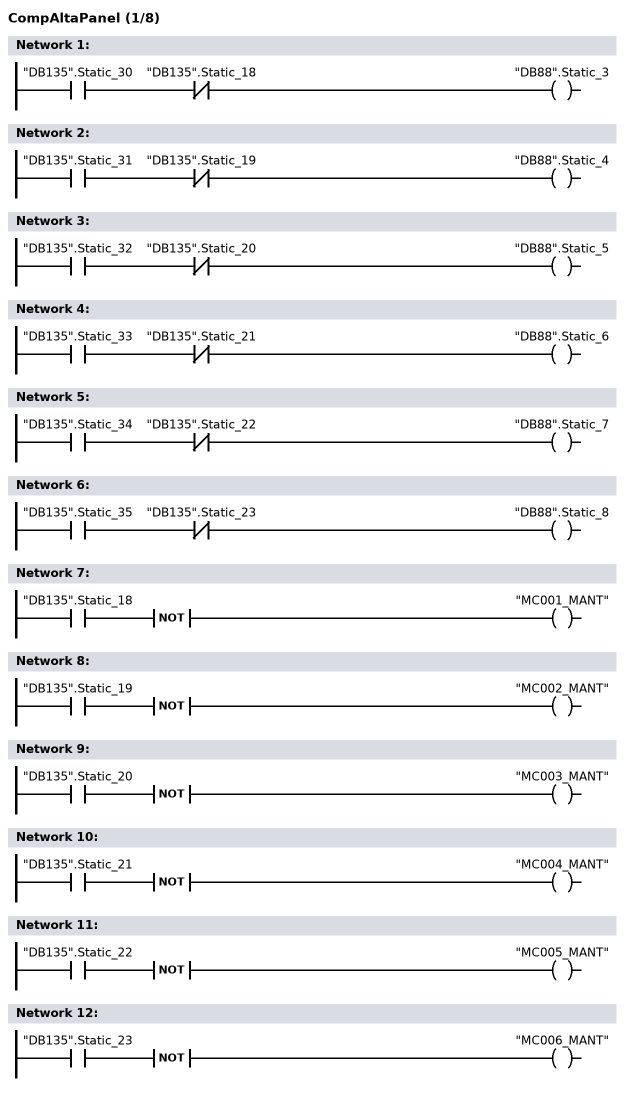
   RUNG wire#powerrail
      Contact( "DB135".Static_30 )
      I_Contact( "DB135".Static_18 )
      Coil( "DB88".Static_3 )
   END_RUNG
   // the same network as SCL:
   "DB88".Static_3 := "DB135".Static_30 AND NOT "DB135".Static_18;
END_REGION

REGION Network 2
   RUNG wire#powerrail
      Contact( "DB135".Static_31 )
      I_Contact( "DB135".Static_19 )
      Coil( "DB88".Static_4 )
   END_RUNG
   // the same network as SCL:
   "DB88".Static_4 := "DB135".Static_31 AND NOT "DB135".Static_19;
END_REGION

REGION Network 3
   RUNG wire#powerrail
      Contact( "DB135".Static_32 )
      I_Contact( "DB135".Static_20 )
      Coil( "DB88".Static_5 )
   END_RUNG
   // the same network as SCL:
   "DB88".Static_5 := "DB135".Static_32 AND NOT "DB135".Static_20;
END_REGION

REGION Network 4
   RUNG wire#powerrail
      Contact( "DB135".Static_33 )
      I_Contact( "DB135".Static_21 )
      Coil( "DB88".Static_6 )
   END_RUNG
   // the same network as SCL:
   "DB88".Static_6 := "DB135".Static_33 AND NOT "DB135".Static_21;
END_REGION

REGION Network 5
   RUNG wire#powerrail
      Contact( "DB135".Static_34 )
      I_Contact( "DB135".Static_22 )
      Coil( "DB88".Static_7 )
   END_RUNG
   // the same network as SCL:
   "DB88".Static_7 := "DB135".Static_34 AND NOT "DB135".Static_22;
END_REGION

REGION Network 6
   RUNG wire#powerrail
      Contact( "DB135".Static_35 )
      I_Contact( "DB135".Static_23 )
      Coil( "DB88".Static_8 )
   END_RUNG
   // the same network as SCL:
   "DB88".Static_8 := "DB135".Static_35 AND NOT "DB135".Static_23;
END_REGION

REGION Network 7
   RUNG wire#powerrail
      Contact( "DB135".Static_18 )
      Not()
      Coil( "MC001_MANT" )
   END_RUNG
   // the same network as SCL:
   "MC001_MANT" := NOT "DB135".Static_18;
END_REGION

REGION Network 8
   RUNG wire#powerrail
      Contact( "DB135".Static_19 )
      Not()
      Coil( "MC002_MANT" )
   END_RUNG
   // the same network as SCL:
   "MC002_MANT" := NOT "DB135".Static_19;
END_REGION

REGION Network 9
   RUNG wire#powerrail
      Contact( "DB135".Static_20 )
      Not()
      Coil( "MC003_MANT" )
   END_RUNG
   // the same network as SCL:
   "MC003_MANT" := NOT "DB135".Static_20;
END_REGION

REGION Network 10
   RUNG wire#powerrail
      Contact( "DB135".Static_21 )
      Not()
      Coil( "MC004_MANT" )
   END_RUNG
   // the same network as SCL:
   "MC004_MANT" := NOT "DB135".Static_21;
END_REGION

REGION Network 11
   RUNG wire#powerrail
      Contact( "DB135".Static_22 )
      Not()
      Coil( "MC005_MANT" )
   END_RUNG
   // the same network as SCL:
   "MC005_MANT" := NOT "DB135".Static_22;
END_REGION

REGION Network 12
   RUNG wire#powerrail
      Contact( "DB135".Static_23 )
      Not()
      Coil( "MC006_MANT" )
   END_RUNG
   // the same network as SCL:
   "MC006_MANT" := NOT "DB135".Static_23;
END_REGION

REGION Network 13
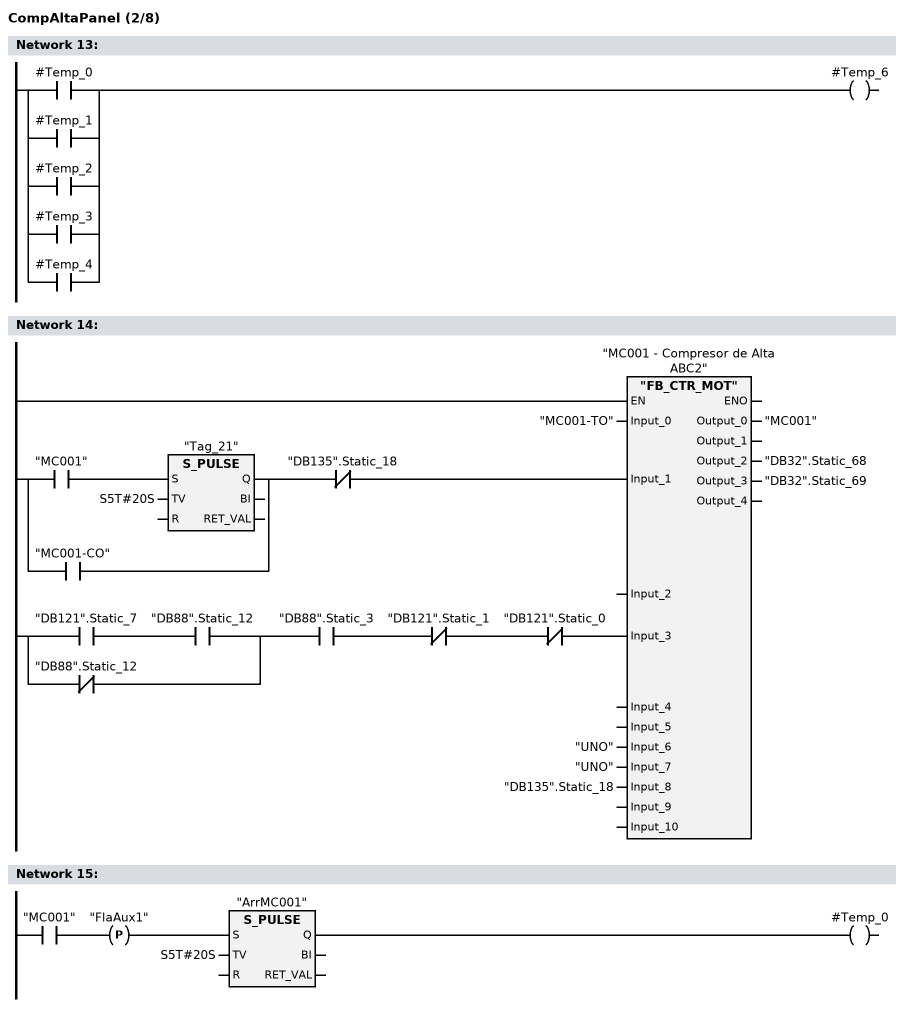
   RUNG wire#powerrail
      Contact( #Temp_0 )
      wire#w1
      Coil( #Temp_6 )
   END_RUNG
   RUNG wire#powerrail
      Contact( #Temp_1 )
   END_RUNG wire#w1
   RUNG wire#powerrail
      Contact( #Temp_2 )
   END_RUNG wire#w1
   RUNG wire#powerrail
      Contact( #Temp_3 )
   END_RUNG wire#w1
   RUNG wire#powerrail
      Contact( #Temp_4 )
   END_RUNG wire#w1
   // the same network as SCL:
   #Temp_6 := #Temp_0 OR #Temp_1 OR #Temp_2 OR #Temp_3 OR #Temp_4;
END_REGION

REGION Network 14
   #_s5time1 := S_PULSE(T_NO := "Tag_21", TV := S5T#20S, S := "MC001", Q => #_w1);
   "MC001 - Compresor de Alta ABC2"(Input_0 := "MC001-TO",   // "FB_CTR_MOT"
                           Input_1 := (#_w1 OR "MC001-CO") AND NOT "DB135".Static_18,
                           Input_3 := (("DB121".Static_7 AND "DB88".Static_12) OR NOT "DB88".Static_12) AND "DB88".Static_3 AND NOT "DB121".Static_1 AND NOT "DB121".Static_0,
                           Input_6 := "UNO",
                           Input_7 := "UNO",
                           Input_8 := "DB135".Static_18,
                           Output_0 => "MC001",
                           Output_2 => "DB32".Static_68,
                           Output_3 => "DB32".Static_69);
END_REGION

REGION Network 15
   RUNG wire#powerrail
      Contact( "MC001" )
      P_Trig( "FlaAux1" )
      S_PULSE(T_NO := "ArrMC001", TV := S5T#20S, R :=, BI =>, RET_VAL =>)
      Coil( #Temp_0 )
   END_RUNG
   // the same network as SCL:
   #_w1 := "MC001" AND NOT "FlaAux1";   // rising edge
   "FlaAux1" := "MC001";
   #_s5time1 := S_PULSE(T_NO := "ArrMC001", S := #_w1, TV := S5T#20S, Q => #_w2);
   #Temp_0 := #_w2;
END_REGION

REGION Network 16
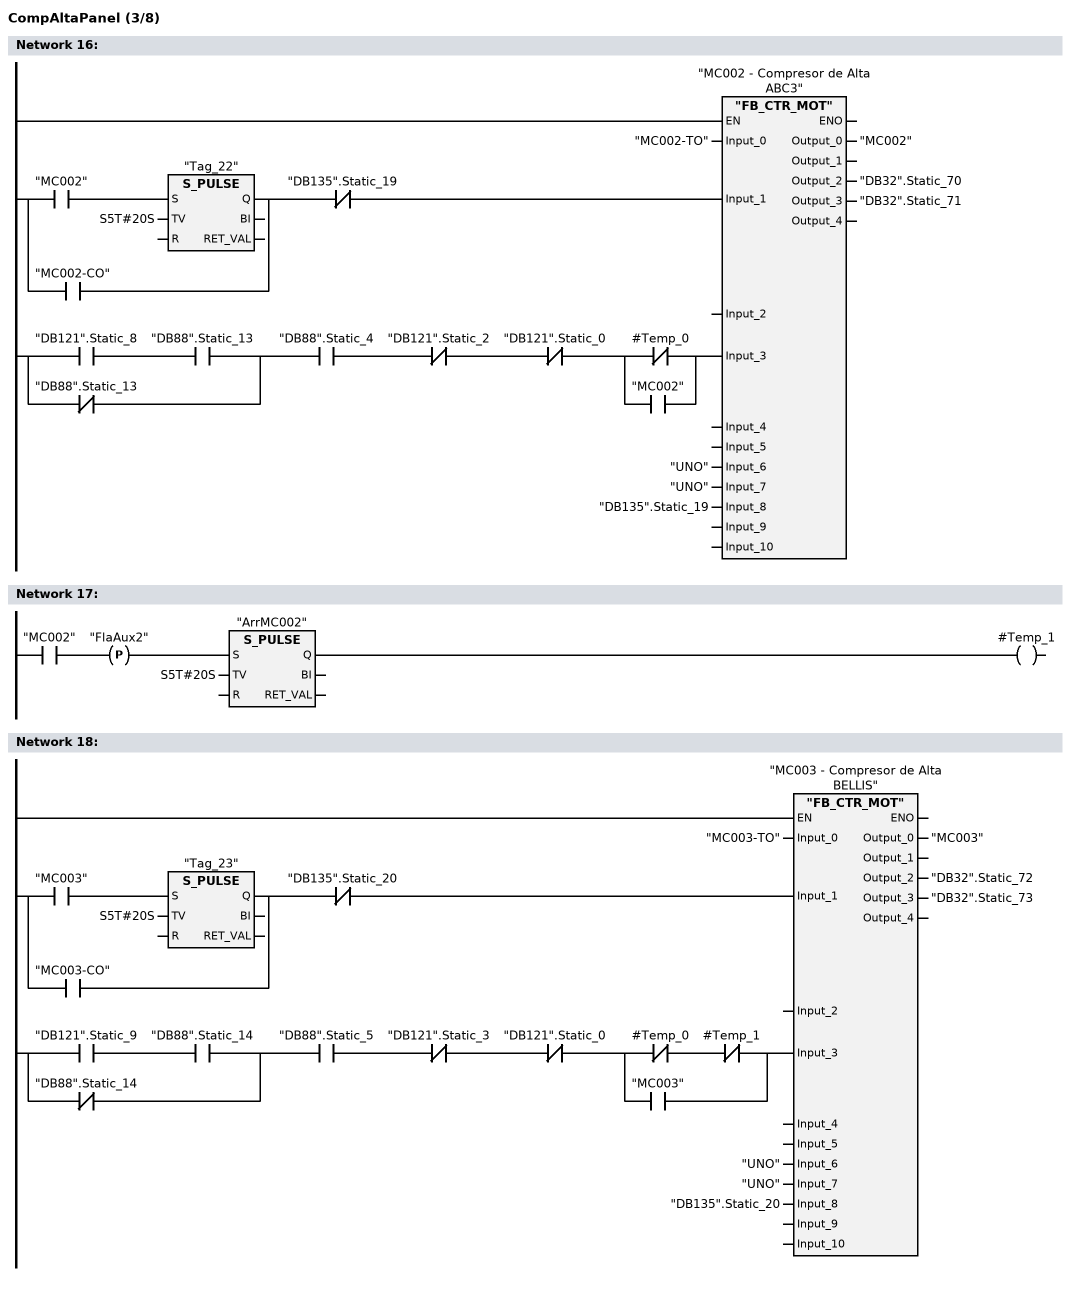
   #_s5time1 := S_PULSE(T_NO := "Tag_22", TV := S5T#20S, S := "MC002", Q => #_w1);
   "MC002 - Compresor de Alta ABC3"(Input_0 := "MC002-TO",   // "FB_CTR_MOT"
                           Input_1 := (#_w1 OR "MC002-CO") AND NOT "DB135".Static_19,
                           Input_3 := (("DB121".Static_8 AND "DB88".Static_13) OR NOT "DB88".Static_13) AND "DB88".Static_4 AND NOT "DB121".Static_2 AND NOT "DB121".Static_0 AND (NOT #Temp_0 OR "MC002"),
                           Input_6 := "UNO",
                           Input_7 := "UNO",
                           Input_8 := "DB135".Static_19,
                           Output_0 => "MC002",
                           Output_2 => "DB32".Static_70,
                           Output_3 => "DB32".Static_71);
END_REGION

REGION Network 17
   RUNG wire#powerrail
      Contact( "MC002" )
      P_Trig( "FlaAux2" )
      S_PULSE(T_NO := "ArrMC002", TV := S5T#20S, R :=, BI =>, RET_VAL =>)
      Coil( #Temp_1 )
   END_RUNG
   // the same network as SCL:
   #_w1 := "MC002" AND NOT "FlaAux2";   // rising edge
   "FlaAux2" := "MC002";
   #_s5time1 := S_PULSE(T_NO := "ArrMC002", S := #_w1, TV := S5T#20S, Q => #_w2);
   #Temp_1 := #_w2;
END_REGION

REGION Network 18
   #_s5time1 := S_PULSE(T_NO := "Tag_23", TV := S5T#20S, S := "MC003", Q => #_w1);
   "MC003 - Compresor de Alta BELLIS"(Input_0 := "MC003-TO",   // "FB_CTR_MOT"
                           Input_1 := (#_w1 OR "MC003-CO") AND NOT "DB135".Static_20,
                           Input_3 := (("DB121".Static_9 AND "DB88".Static_14) OR NOT "DB88".Static_14) AND "DB88".Static_5 AND NOT "DB121".Static_3 AND NOT "DB121".Static_0 AND ((NOT #Temp_0 AND NOT #Temp_1) OR "MC003"),
                           Input_6 := "UNO",
                           Input_7 := "UNO",
                           Input_8 := "DB135".Static_20,
                           Output_0 => "MC003",
                           Output_2 => "DB32".Static_72,
                           Output_3 => "DB32".Static_73);
END_REGION

REGION Network 19
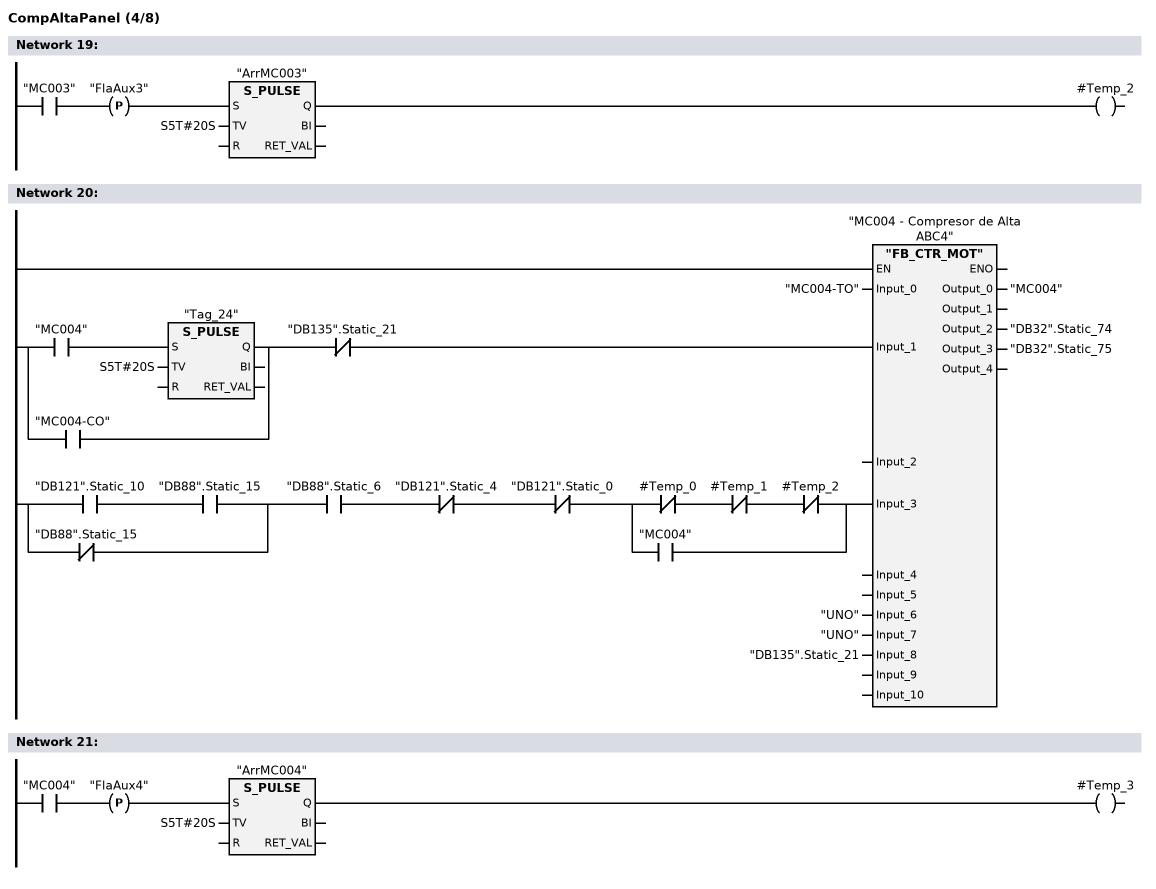
   RUNG wire#powerrail
      Contact( "MC003" )
      P_Trig( "FlaAux3" )
      S_PULSE(T_NO := "ArrMC003", TV := S5T#20S, R :=, BI =>, RET_VAL =>)
      Coil( #Temp_2 )
   END_RUNG
   // the same network as SCL:
   #_w1 := "MC003" AND NOT "FlaAux3";   // rising edge
   "FlaAux3" := "MC003";
   #_s5time1 := S_PULSE(T_NO := "ArrMC003", S := #_w1, TV := S5T#20S, Q => #_w2);
   #Temp_2 := #_w2;
END_REGION

REGION Network 20
   #_s5time1 := S_PULSE(T_NO := "Tag_24", TV := S5T#20S, S := "MC004", Q => #_w1);
   "MC004 - Compresor de Alta ABC4"(Input_0 := "MC004-TO",   // "FB_CTR_MOT"
                           Input_1 := (#_w1 OR "MC004-CO") AND NOT "DB135".Static_21,
                           Input_3 := (("DB121".Static_10 AND "DB88".Static_15) OR NOT "DB88".Static_15) AND "DB88".Static_6 AND NOT "DB121".Static_4 AND NOT "DB121".Static_0 AND ((NOT #Temp_0 AND NOT #Temp_1 AND NOT #Temp_2) OR "MC004"),
                           Input_6 := "UNO",
                           Input_7 := "UNO",
                           Input_8 := "DB135".Static_21,
                           Output_0 => "MC004",
                           Output_2 => "DB32".Static_74,
                           Output_3 => "DB32".Static_75);
END_REGION

REGION Network 21
   RUNG wire#powerrail
      Contact( "MC004" )
      P_Trig( "FlaAux4" )
      S_PULSE(T_NO := "ArrMC004", TV := S5T#20S, R :=, BI =>, RET_VAL =>)
      Coil( #Temp_3 )
   END_RUNG
   // the same network as SCL:
   #_w1 := "MC004" AND NOT "FlaAux4";   // rising edge
   "FlaAux4" := "MC004";
   #_s5time1 := S_PULSE(T_NO := "ArrMC004", S := #_w1, TV := S5T#20S, Q => #_w2);
   #Temp_3 := #_w2;
END_REGION

REGION Network 22
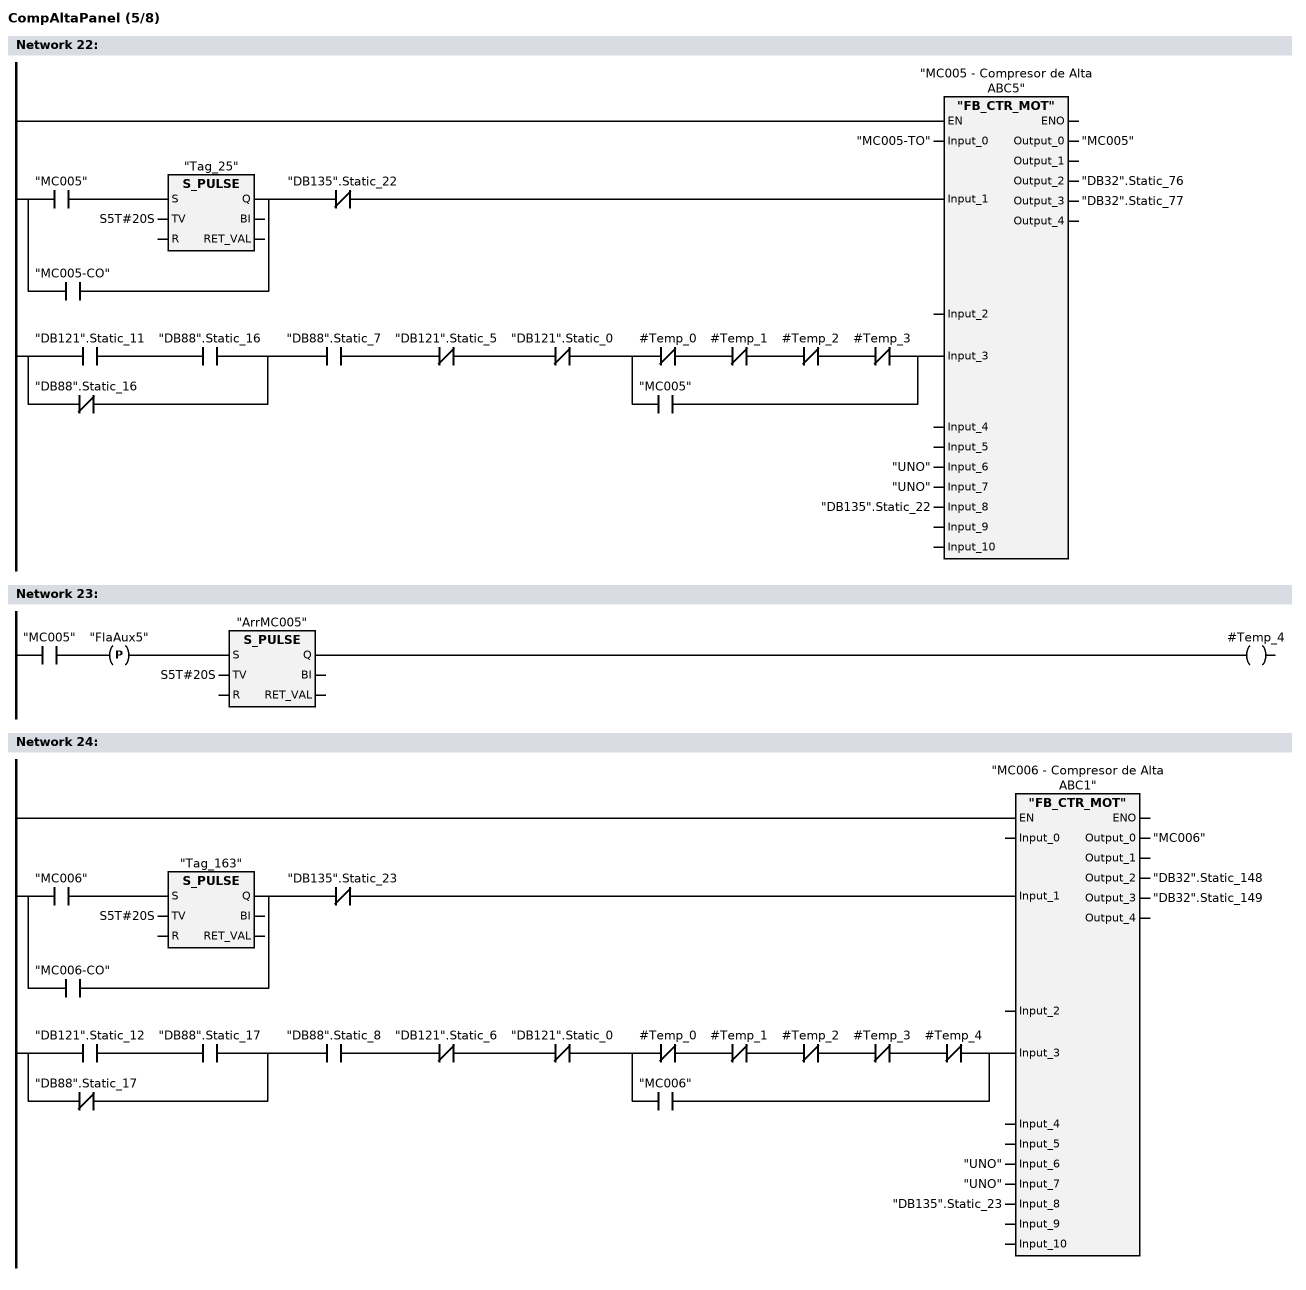
   #_s5time1 := S_PULSE(T_NO := "Tag_25", TV := S5T#20S, S := "MC005", Q => #_w1);
   "MC005 - Compresor de Alta ABC5"(Input_0 := "MC005-TO",   // "FB_CTR_MOT"
                           Input_1 := (#_w1 OR "MC005-CO") AND NOT "DB135".Static_22,
                           Input_3 := (("DB121".Static_11 AND "DB88".Static_16) OR NOT "DB88".Static_16) AND "DB88".Static_7 AND NOT "DB121".Static_5 AND NOT "DB121".Static_0 AND ((NOT #Temp_0 AND NOT #Temp_1 AND NOT #Temp_2 AND NOT #Temp_3) OR "MC005"),
                           Input_6 := "UNO",
                           Input_7 := "UNO",
                           Input_8 := "DB135".Static_22,
                           Output_0 => "MC005",
                           Output_2 => "DB32".Static_76,
                           Output_3 => "DB32".Static_77);
END_REGION

REGION Network 23
   RUNG wire#powerrail
      Contact( "MC005" )
      P_Trig( "FlaAux5" )
      S_PULSE(T_NO := "ArrMC005", TV := S5T#20S, R :=, BI =>, RET_VAL =>)
      Coil( #Temp_4 )
   END_RUNG
   // the same network as SCL:
   #_w1 := "MC005" AND NOT "FlaAux5";   // rising edge
   "FlaAux5" := "MC005";
   #_s5time1 := S_PULSE(T_NO := "ArrMC005", S := #_w1, TV := S5T#20S, Q => #_w2);
   #Temp_4 := #_w2;
END_REGION

REGION Network 24
   #_s5time1 := S_PULSE(T_NO := "Tag_163", TV := S5T#20S, S := "MC006", Q => #_w1);
   "MC006 - Compresor de Alta ABC1"(Input_1 := (#_w1 OR "MC006-CO") AND NOT "DB135".Static_23,   // "FB_CTR_MOT"
                           Input_3 := (("DB121".Static_12 AND "DB88".Static_17) OR NOT "DB88".Static_17) AND "DB88".Static_8 AND NOT "DB121".Static_6 AND NOT "DB121".Static_0 AND ((NOT #Temp_0 AND NOT #Temp_1 AND NOT #Temp_2 AND NOT #Temp_3 AND NOT #Temp_4) OR "MC006"),
                           Input_6 := "UNO",
                           Input_7 := "UNO",
                           Input_8 := "DB135".Static_23,
                           Output_0 => "MC006",
                           Output_2 => "DB32".Static_148,
                           Output_3 => "DB32".Static_149);
END_REGION

REGION Network 25
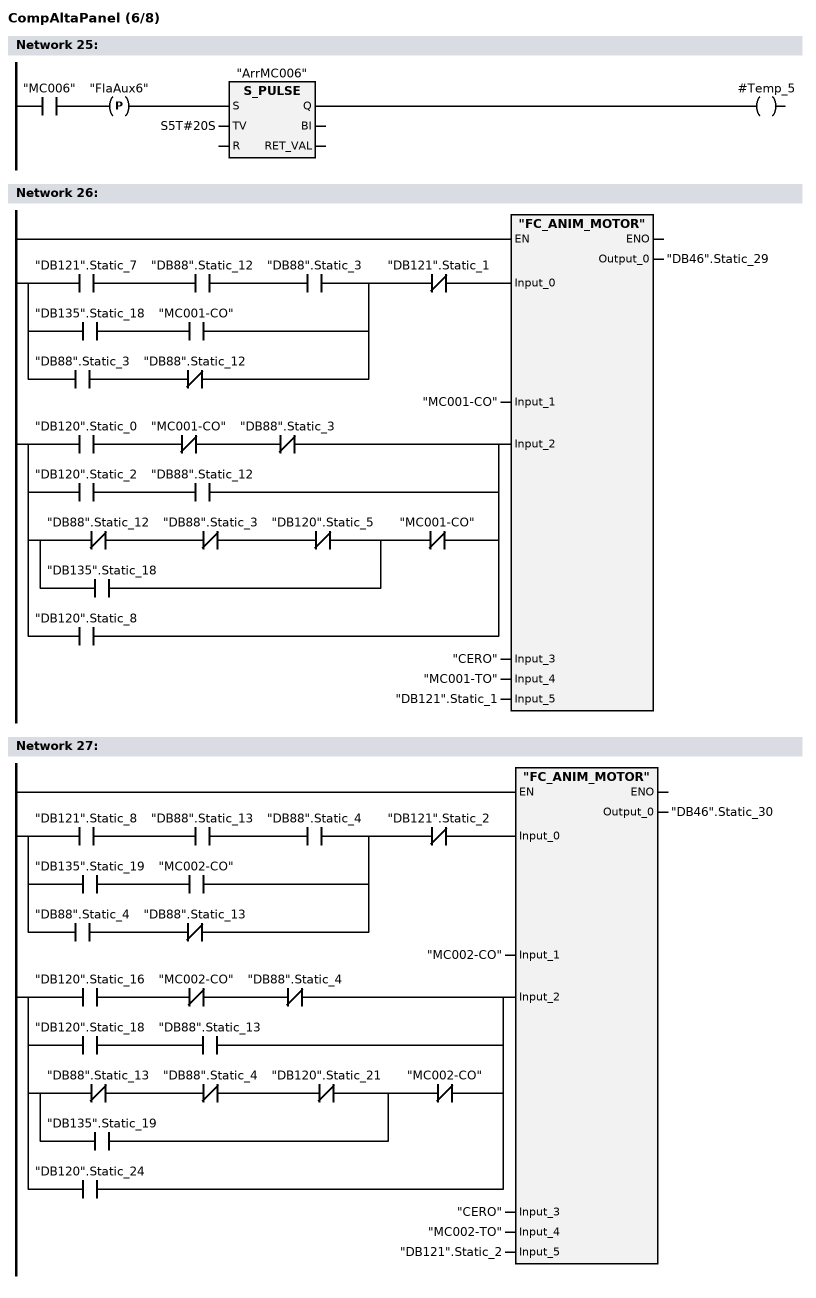
   RUNG wire#powerrail
      Contact( "MC006" )
      P_Trig( "FlaAux6" )
      S_PULSE(T_NO := "ArrMC006", TV := S5T#20S, R :=, BI =>, RET_VAL =>)
      Coil( #Temp_5 )
   END_RUNG
   // the same network as SCL:
   #_w1 := "MC006" AND NOT "FlaAux6";   // rising edge
   "FlaAux6" := "MC006";
   #_s5time1 := S_PULSE(T_NO := "ArrMC006", S := #_w1, TV := S5T#20S, Q => #_w2);
   #Temp_5 := #_w2;
END_REGION

REGION Network 26
   "FC_ANIM_MOTOR"(Input_0 := (("DB121".Static_7 AND "DB88".Static_12 AND "DB88".Static_3) OR ("DB135".Static_18 AND "MC001-CO") OR ("DB88".Static_3 AND NOT "DB88".Static_12)) AND NOT "DB121".Static_1,
                   Input_1 := "MC001-CO",
                   Input_2 := ("DB120".Static_0 AND NOT "MC001-CO" AND NOT "DB88".Static_3) OR ("DB120".Static_2 AND "DB88".Static_12) OR "DB120".Static_8 OR (("DB135".Static_18 OR (NOT "DB88".Static_12 AND NOT "DB88".Static_3 AND NOT "DB120".Static_5)) AND NOT "MC001-CO"),
                   Input_3 := "CERO",
                   Input_4 := "MC001-TO",
                   Input_5 := "DB121".Static_1,
                   Output_0 => "DB46".Static_29);
END_REGION

REGION Network 27
   "FC_ANIM_MOTOR"(Input_0 := (("DB121".Static_8 AND "DB88".Static_13 AND "DB88".Static_4) OR ("DB135".Static_19 AND "MC002-CO") OR ("DB88".Static_4 AND NOT "DB88".Static_13)) AND NOT "DB121".Static_2,
                   Input_1 := "MC002-CO",
                   Input_2 := ("DB120".Static_16 AND NOT "MC002-CO" AND NOT "DB88".Static_4) OR ("DB120".Static_18 AND "DB88".Static_13) OR "DB120".Static_24 OR (("DB135".Static_19 OR (NOT "DB88".Static_13 AND NOT "DB88".Static_4 AND NOT "DB120".Static_21)) AND NOT "MC002-CO"),
                   Input_3 := "CERO",
                   Input_4 := "MC002-TO",
                   Input_5 := "DB121".Static_2,
                   Output_0 => "DB46".Static_30);
END_REGION

REGION Network 28
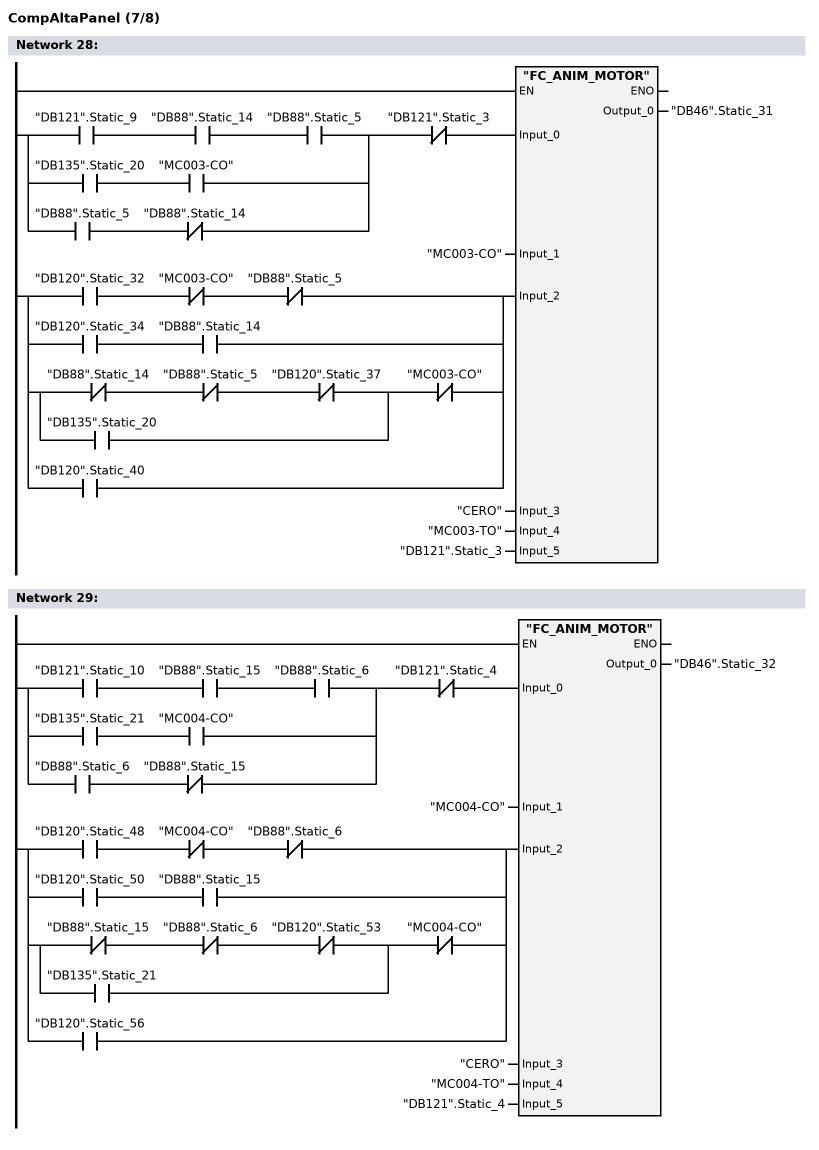
   "FC_ANIM_MOTOR"(Input_0 := (("DB121".Static_9 AND "DB88".Static_14 AND "DB88".Static_5) OR ("DB135".Static_20 AND "MC003-CO") OR ("DB88".Static_5 AND NOT "DB88".Static_14)) AND NOT "DB121".Static_3,
                   Input_1 := "MC003-CO",
                   Input_2 := ("DB120".Static_32 AND NOT "MC003-CO" AND NOT "DB88".Static_5) OR ("DB120".Static_34 AND "DB88".Static_14) OR "DB120".Static_40 OR (("DB135".Static_20 OR (NOT "DB88".Static_14 AND NOT "DB88".Static_5 AND NOT "DB120".Static_37)) AND NOT "MC003-CO"),
                   Input_3 := "CERO",
                   Input_4 := "MC003-TO",
                   Input_5 := "DB121".Static_3,
                   Output_0 => "DB46".Static_31);
END_REGION

REGION Network 29
   "FC_ANIM_MOTOR"(Input_0 := (("DB121".Static_10 AND "DB88".Static_15 AND "DB88".Static_6) OR ("DB135".Static_21 AND "MC004-CO") OR ("DB88".Static_6 AND NOT "DB88".Static_15)) AND NOT "DB121".Static_4,
                   Input_1 := "MC004-CO",
                   Input_2 := ("DB120".Static_48 AND NOT "MC004-CO" AND NOT "DB88".Static_6) OR ("DB120".Static_50 AND "DB88".Static_15) OR "DB120".Static_56 OR (("DB135".Static_21 OR (NOT "DB88".Static_15 AND NOT "DB88".Static_6 AND NOT "DB120".Static_53)) AND NOT "MC004-CO"),
                   Input_3 := "CERO",
                   Input_4 := "MC004-TO",
                   Input_5 := "DB121".Static_4,
                   Output_0 => "DB46".Static_32);
END_REGION

REGION Network 30
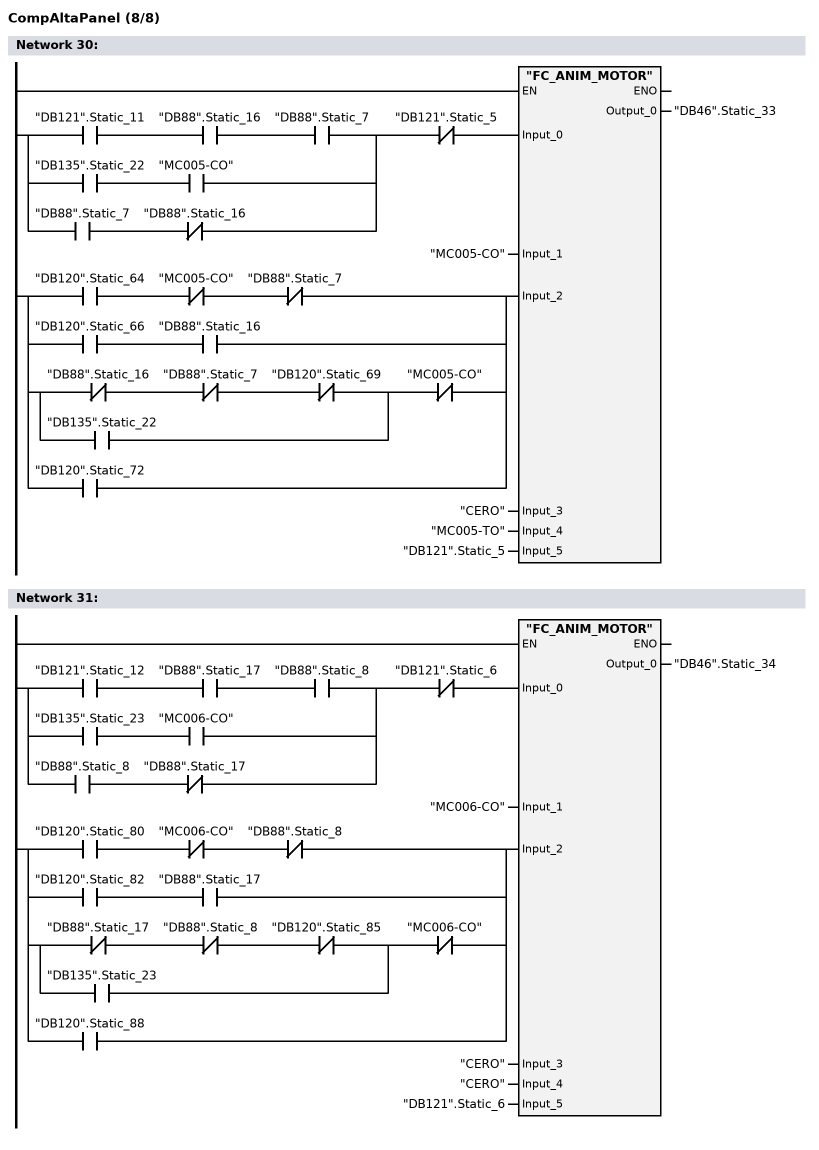
   "FC_ANIM_MOTOR"(Input_0 := (("DB121".Static_11 AND "DB88".Static_16 AND "DB88".Static_7) OR ("DB135".Static_22 AND "MC005-CO") OR ("DB88".Static_7 AND NOT "DB88".Static_16)) AND NOT "DB121".Static_5,
                   Input_1 := "MC005-CO",
                   Input_2 := ("DB120".Static_64 AND NOT "MC005-CO" AND NOT "DB88".Static_7) OR ("DB120".Static_66 AND "DB88".Static_16) OR "DB120".Static_72 OR (("DB135".Static_22 OR (NOT "DB88".Static_16 AND NOT "DB88".Static_7 AND NOT "DB120".Static_69)) AND NOT "MC005-CO"),
                   Input_3 := "CERO",
                   Input_4 := "MC005-TO",
                   Input_5 := "DB121".Static_5,
                   Output_0 => "DB46".Static_33);
END_REGION

REGION Network 31
   "FC_ANIM_MOTOR"(Input_0 := (("DB121".Static_12 AND "DB88".Static_17 AND "DB88".Static_8) OR ("DB135".Static_23 AND "MC006-CO") OR ("DB88".Static_8 AND NOT "DB88".Static_17)) AND NOT "DB121".Static_6,
                   Input_1 := "MC006-CO",
                   Input_2 := ("DB120".Static_80 AND NOT "MC006-CO" AND NOT "DB88".Static_8) OR ("DB120".Static_82 AND "DB88".Static_17) OR "DB120".Static_88 OR (("DB135".Static_23 OR (NOT "DB88".Static_17 AND NOT "DB88".Static_8 AND NOT "DB120".Static_85)) AND NOT "MC006-CO"),
                   Input_3 := "CERO",
                   Input_4 := "CERO",
                   Input_5 := "DB121".Static_6,
                   Output_0 => "DB46".Static_34);
END_REGION
END_FUNCTION

FUNCTION "ModoManualAlta" : Void   // FC48, LAD
{ S7_Optimized_Access := 'FALSE' }
VERSION : 0.1
   VAR_TEMP   // added for the SCL form of the ladder/FBD networks
      _w1 : Bool;
      _s5time1 : S5Time;
   END_VAR
BEGIN

REGION Network 1
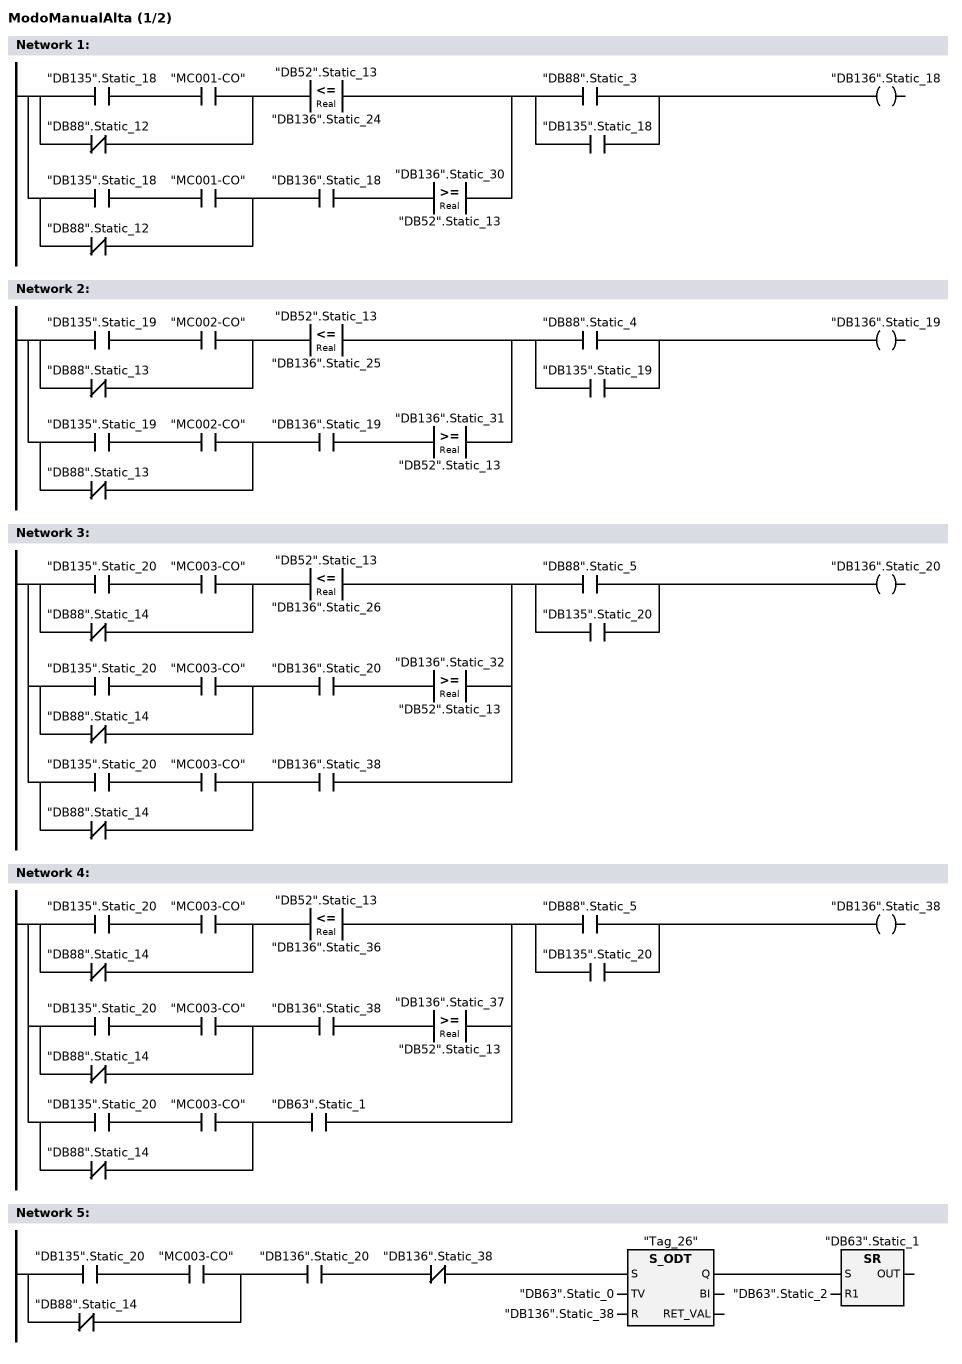
   "DB136".Static_18 := (((NOT "DB88".Static_12 OR ("DB135".Static_18 AND "MC001-CO")) AND ("DB52".Static_13 <= "DB136".Static_24)) OR ((NOT "DB88".Static_12 OR ("DB135".Static_18 AND "MC001-CO")) AND "DB136".Static_18 AND ("DB136".Static_30 >= "DB52".Static_13))) AND ("DB88".Static_3 OR "DB135".Static_18);
END_REGION

REGION Network 2
   "DB136".Static_19 := (((NOT "DB88".Static_13 OR ("DB135".Static_19 AND "MC002-CO")) AND ("DB52".Static_13 <= "DB136".Static_25)) OR ((NOT "DB88".Static_13 OR ("DB135".Static_19 AND "MC002-CO")) AND "DB136".Static_19 AND ("DB136".Static_31 >= "DB52".Static_13))) AND ("DB88".Static_4 OR "DB135".Static_19);
END_REGION

REGION Network 3
   "DB136".Static_20 := (((NOT "DB88".Static_14 OR ("DB135".Static_20 AND "MC003-CO")) AND ("DB52".Static_13 <= "DB136".Static_26)) OR ((NOT "DB88".Static_14 OR ("DB135".Static_20 AND "MC003-CO")) AND "DB136".Static_20 AND ("DB136".Static_32 >= "DB52".Static_13)) OR ((NOT "DB88".Static_14 OR ("DB135".Static_20 AND "MC003-CO")) AND "DB136".Static_38)) AND ("DB88".Static_5 OR "DB135".Static_20);
END_REGION

REGION Network 4
   "DB136".Static_38 := (((NOT "DB88".Static_14 OR ("DB135".Static_20 AND "MC003-CO")) AND ("DB52".Static_13 <= "DB136".Static_36)) OR ((NOT "DB88".Static_14 OR ("DB135".Static_20 AND "MC003-CO")) AND "DB136".Static_38 AND ("DB136".Static_37 >= "DB52".Static_13)) OR ((NOT "DB88".Static_14 OR ("DB135".Static_20 AND "MC003-CO")) AND "DB63".Static_1)) AND ("DB88".Static_5 OR "DB135".Static_20);
END_REGION

REGION Network 5
   #_s5time1 := S_ODT(T_NO := "Tag_26",
                      TV := "DB63".Static_0,
                      R := "DB136".Static_38,
                      S := (NOT "DB88".Static_14 OR ("DB135".Static_20 AND "MC003-CO")) AND "DB136".Static_20 AND NOT "DB136".Static_38,
                      Q => #_w1);
   IF #_w1 THEN
       "DB63".Static_1 := TRUE;   // SR flip-flop
   END_IF;
   IF "DB63".Static_2 THEN "DB63".Static_1 := FALSE; END_IF;
END_REGION

REGION Network 6